(* Logix 5000 project; controller _GigaDiscovery vendor 1 type 14 code 244 rev 35.11; software revision 35.03; part 9 of 23 *)
(* tags used below, declared in another part *)
   Pylon_Sequencer : Sequencer;
   Acc_Time : REAL;   // T2 Region 2
   Auto_Cycle_Step : DINT;
   Automatic_Cycle_DB : Auto_Cycle[6];
   Cycle_Time : TIMER;
   Direction : BOOL;   // 1 = Spinta CW 0 = Spinta CCW
   Echo_HMI_Modify_Auto_Cycle_Ptr : DINT;
   Emergencies_CL1 : DINT[14];
   Gondola_Speed_Reference : DINT;
   HMI_Auto_Cycle_in_Modify : Auto_Cycle;
   HMI_Auto_Cycle_Step_Modify : DINT;
   HMI_Modify_Auto_Cycle_Ptr : DINT;
   HMI_Save_Recipe : BOOL;
   HMI_Step_in_Modify_Gondola_Speed : DINT;
   HMI_Step_in_Modify_Gondola_Time : DINT;
   HMI_Work_Auto_Cycle_Ptr : DINT;
   Jerk_Time : REAL;   // T1 Region 1
   K_Inversion : REAL;   // Fattore di Inversione
   K_Inversion_SCRV : REAL;
   LapBarsMonitor : LapBars_Monitor[41];
   LPF_WLang_Speed_to_Torq : REAL;
   ONP : DINT;   // Optional Not Present
   Oscillation_Error : REAL;
   PW_Bool : BOOL[32];
   PW_Dint : DINT[64];
   Pylon_Axe : Axe;
   Pylon_Filtered_Speed : REAL;
   RESTRAINTS_Open_Postion : BOOL[64];
   RESTRAINTS_Sector : LapBars_Sector[9];
   SCuve_K_Stop : S_Curve_Calc;
   Second_Oscillation_Done : BOOL;   // Second Oscillation End
   Start_Stop_Cycle : Sequencer;
   Stop_K_to_Zero : BOOL;
   Target_Angle : REAL;
   To_Sfty : Std_to_Sfty;
   Torque_Cmd_from_Cycle : REAL;
   TorquePos_Angle_Control : REAL;
   Work_Auto_Cycle : Auto_Cycle;
   Work_Auto_Cycle_Ptr : DINT;
(* Pylon, continued *)

ROUTINE Main   (* ladder *)
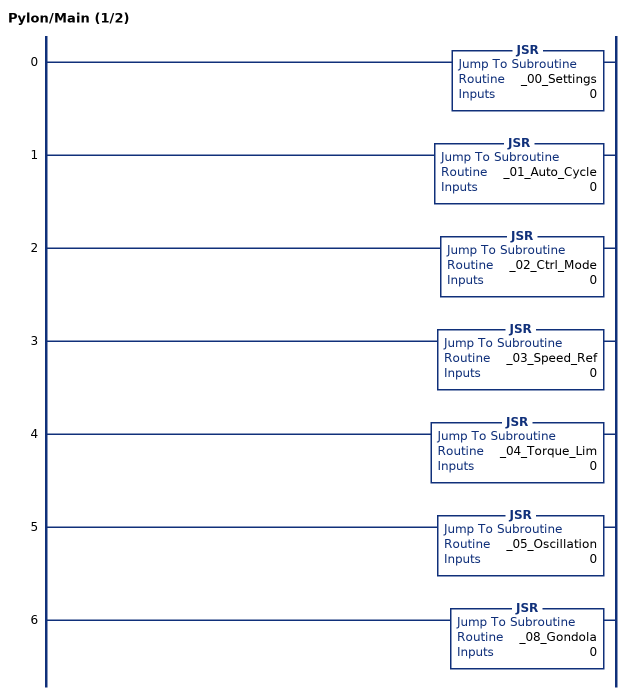
   0: JSR(_00_Settings,0);
   1: JSR(_01_Auto_Cycle,0);
   2: JSR(_02_Ctrl_Mode,0);
   3: JSR(_03_Speed_Ref,0);
   4: JSR(_04_Torque_Lim,0);
   5: JSR(_05_Oscillation,0);
   6: JSR(_08_Gondola,0);
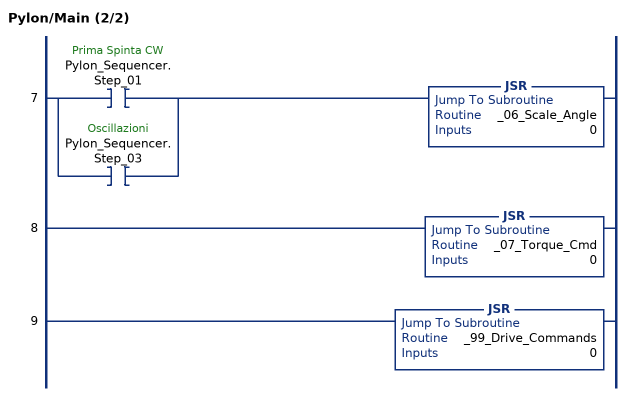
   7: [XIC(Pylon_Sequencer.Step_01) ,XIC(Pylon_Sequencer.Step_03) ]JSR(_06_Scale_Angle,0);
   8: JSR(_07_Torque_Cmd,0);
   9: JSR(_99_Drive_Commands,0);
END_ROUTINE
END_PROGRAM

PROGRAM Pylon_Oscillation   (* main routine _00_Oscillation *)
VAR
   ADD_01 : FBD_MATH := (SourceA := 0.3, SourceB := 0.5, Dest := 0.8);
   BOR_01 : FBD_BOOLEAN_OR;
   DIV_01 : FBD_MATH := (SourceA := 86.0, SourceB := 0.8, Dest := 107.5);
   DIV_02 : FBD_MATH := (SourceA := 107.5, SourceB := 0.3, Dest := 358.3333);
   GRT_01 : FBD_COMPARE;
   LES_01 : FBD_COMPARE;
   NEG_01 : FBD_MATH_ADVANCED := (Source := 77.39982, Dest := -77.39982);
   OSRI_01 : FBD_ONESHOT;
   OSRI_02 : FBD_ONESHOT;
   SCRV_01 : S_CURVE := (AccelRate := 107.5, DecelRate := 107.5, JerkRate := 358.3333, RTSTime := 1, DeltaT := 0.005);
   SCRV_02 : S_CURVE := (In := -10.0, AccelRate := 25.0, DecelRate := 25.0, JerkRate := 25.0, RTSTime := 1, Out := -10.0, DeltaT := 0.005);
   SEL_01 : SELECT := (In1 := 119.95556, In2 := 119.95556, Out := 119.95556);
   SUB_02 : FBD_MATH := (SourceA := 120.0, SourceB := 0.044444446, Dest := 119.95556);
END_VAR

ROUTINE _00_Oscillation   (* function block diagram *)
   SHEET 1
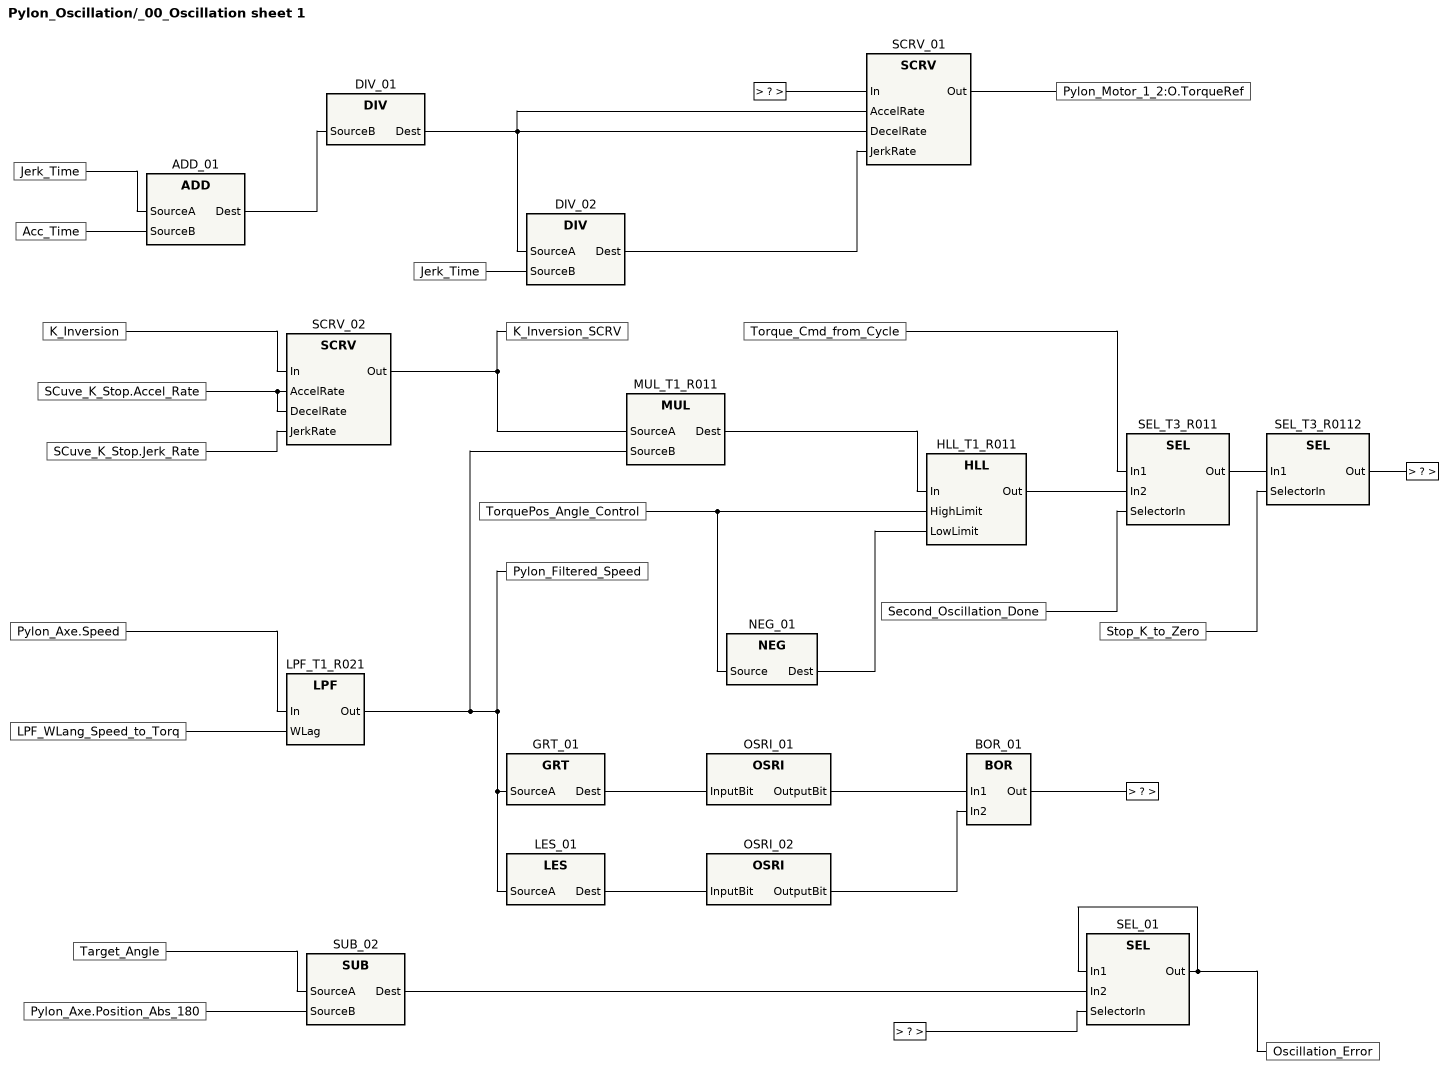
   ADD_01 : ADD(SourceA := Jerk_Time, SourceB := Acc_Time);
   SCRV_02 : SCRV(In := K_Inversion, AccelRate := SCuve_K_Stop.Accel_Rate, DecelRate := SCuve_K_Stop.Accel_Rate, JerkRate := SCuve_K_Stop.Jerk_Rate);
   LPF_T1_R021 : LPF(In := Pylon_Axe.Speed, WLag := LPF_WLang_Speed_to_Torq);
   SUB_02 : SUB(SourceA := Target_Angle, SourceB := Pylon_Axe.Position_Abs_180);
   DIV_01 : DIV(SourceB := ADD_01.Dest);
   K_Inversion_SCRV := SCRV_02.Out;
   Pylon_Filtered_Speed := LPF_T1_R021.Out;
   GRT_01 : GRT(SourceA := LPF_T1_R021.Out);
   LES_01 : LES(SourceA := LPF_T1_R021.Out);
   DIV_02 : DIV(SourceA := DIV_01.Dest, SourceB := Jerk_Time);
   MUL_T1_R011 : MUL(SourceA := SCRV_02.Out, SourceB := LPF_T1_R021.Out);
   OSRI_01 : OSRI(InputBit := GRT_01.Dest);
   OSRI_02 : OSRI(InputBit := LES_01.Dest);
   NEG_01 : NEG(Source := TorquePos_Angle_Control);
   HLL_T1_R011 : HLL(In := MUL_T1_R011.Dest, HighLimit := TorquePos_Angle_Control, LowLimit := NEG_01.Dest);
   BOR_01 : BOR(In1 := OSRI_01.OutputBit, In2 := OSRI_02.OutputBit);
   SEL_T3_R011 : SEL(In1 := Torque_Cmd_from_Cycle, In2 := HLL_T1_R011.Out, SelectorIn := Second_Oscillation_Done);
   WIRE(?) := BOR_01.Out;
   SEL_T3_R0112 : SEL(In1 := SEL_T3_R011.Out, SelectorIn := Stop_K_to_Zero);
   WIRE(?) := SEL_T3_R0112.Out;
   SCRV_01 : SCRV(In := WIRE(?), AccelRate := DIV_01.Dest, DecelRate := DIV_01.Dest, JerkRate := DIV_02.Dest);
   Pylon_Motor_1_2:O.TorqueRef := SCRV_01.Out;
   SEL_01 : SEL(In1 := SEL_01.Out, In2 := SUB_02.Dest, SelectorIn := WIRE(?));
   Oscillation_Error := SEL_01.Out;
END_ROUTINE
END_PROGRAM

PROGRAM Recipe   (* main routine Main *)
VAR
   Echo_HMI_Auto_Cycle_Step_Modify : DINT := 2;
   HMI_Cycle_Time_to_End : DINT := 145;
   Os : DINT;
   Step_Timer : TIMER := (PRE := 60000);
END_VAR

ROUTINE _01_Auto_Cycle   (* ladder *)
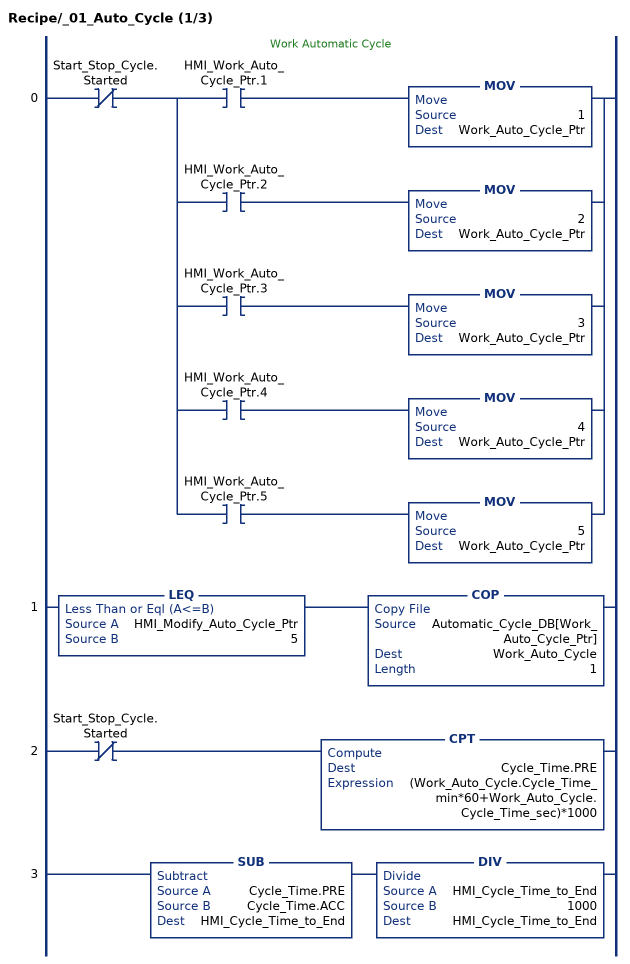
   // Work Automatic Cycle
   0: XIO(Start_Stop_Cycle.Started)[XIC(HMI_Work_Auto_Cycle_Ptr.1) MOV(1,Work_Auto_Cycle_Ptr) ,XIC(HMI_Work_Auto_Cycle_Ptr.2) MOV(2,Work_Auto_Cycle_Ptr) ,XIC(HMI_Work_Auto_Cycle_Ptr.3) MOV(3,Work_Auto_Cycle_Ptr) ,XIC(HMI_Work_Auto_Cycle_Ptr.4) MOV(4,Work_Auto_Cycle_Ptr) ,XIC(HMI_Work_Auto_Cycle_Ptr.5) MOV(5,Work_Auto_Cycle_Ptr) ];
   1: LEQ(HMI_Modify_Auto_Cycle_Ptr,5)COP(Automatic_Cycle_DB[Work_Auto_Cycle_Ptr],Work_Auto_Cycle,1);
   2: XIO(Start_Stop_Cycle.Started)CPT(Cycle_Time.PRE,(Work_Auto_Cycle.Cycle_Time_min*60+Work_Auto_Cycle.Cycle_Time_sec)*1000);
   3: SUB(Cycle_Time.PRE,Cycle_Time.ACC,HMI_Cycle_Time_to_End)DIV(HMI_Cycle_Time_to_End,1000,HMI_Cycle_Time_to_End);
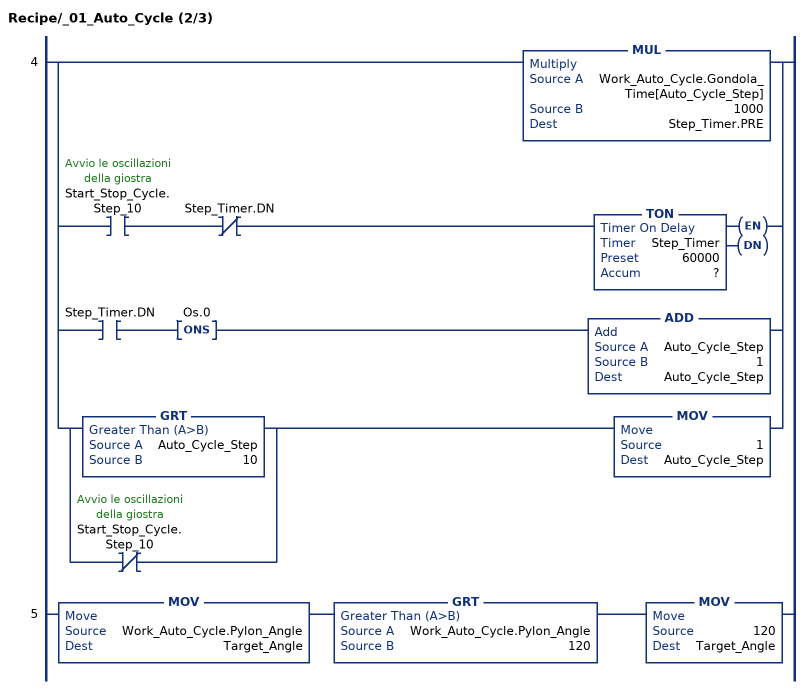
   4: [MUL(Work_Auto_Cycle.Gondola_Time[Auto_Cycle_Step],1000,Step_Timer.PRE) ,XIC(Start_Stop_Cycle.Step_10) XIO(Step_Timer.DN) TON(Step_Timer,?,?) ,XIC(Step_Timer.DN) ONS(Os.0) ADD(Auto_Cycle_Step,1,Auto_Cycle_Step) ,[GRT(Auto_Cycle_Step,10) ,XIO(Start_Stop_Cycle.Step_10) ] MOV(1,Auto_Cycle_Step) ];
   5: MOV(Work_Auto_Cycle.Pylon_Angle,Target_Angle)GRT(Work_Auto_Cycle.Pylon_Angle,120)MOV(120,Target_Angle);
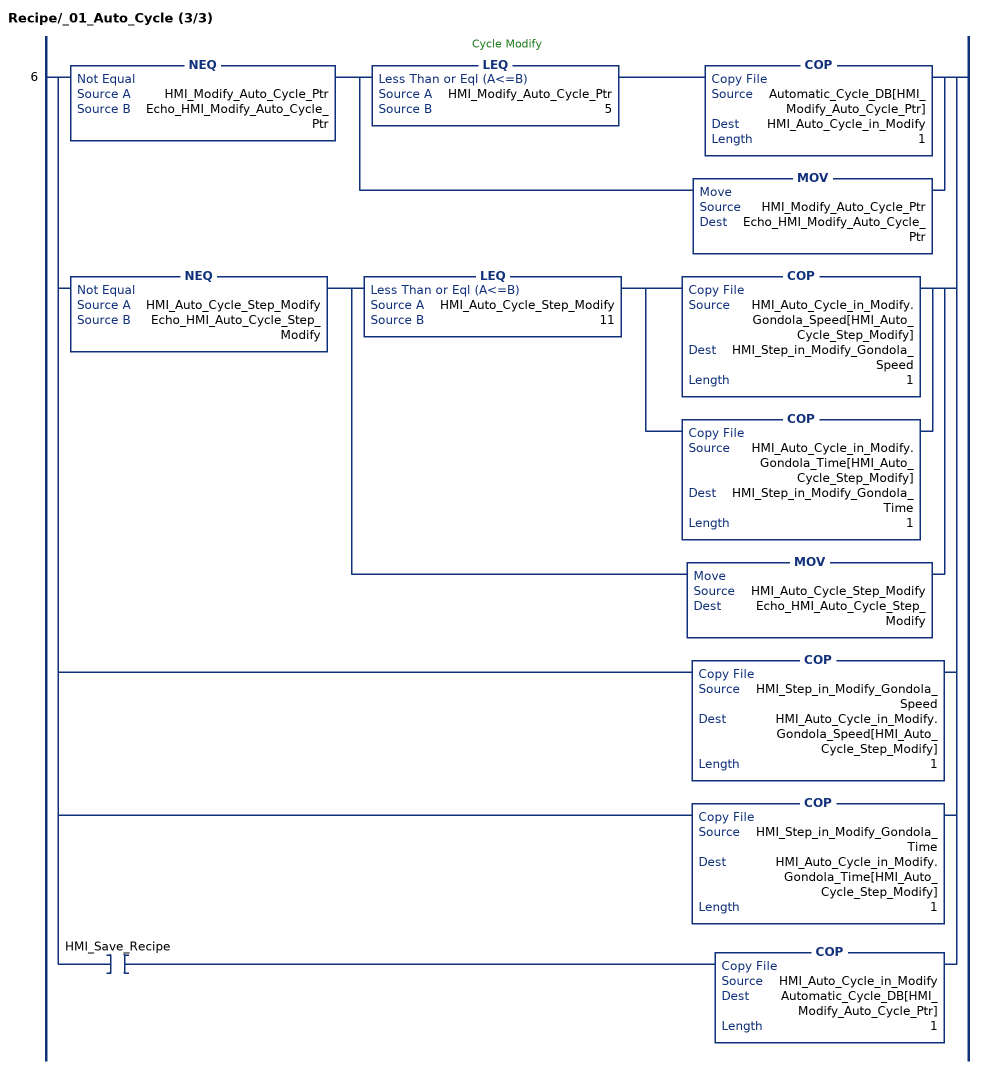
   // Cycle Modify
   6: [NEQ(HMI_Modify_Auto_Cycle_Ptr,Echo_HMI_Modify_Auto_Cycle_Ptr) [LEQ(HMI_Modify_Auto_Cycle_Ptr,5) COP(Automatic_Cycle_DB[HMI_Modify_Auto_Cycle_Ptr],HMI_Auto_Cycle_in_Modify,1) ,MOV(HMI_Modify_Auto_Cycle_Ptr,Echo_HMI_Modify_Auto_Cycle_Ptr) ] ,NEQ(HMI_Auto_Cycle_Step_Modify,Echo_HMI_Auto_Cycle_Step_Modify) [LEQ(HMI_Auto_Cycle_Step_Modify,11) [COP(HMI_Auto_Cycle_in_Modify.Gondola_Speed[HMI_Auto_Cycle_Step_Modify],HMI_Step_in_Modify_Gondola_Speed,1) ,COP(HMI_Auto_Cycle_in_Modify.Gondola_Time[HMI_Auto_Cycle_Step_Modify],HMI_Step_in_Modify_Gondola_Time,1) ] ,MOV(HMI_Auto_Cycle_Step_Modify,Echo_HMI_Auto_Cycle_Step_Modify) ] ,[COP(HMI_Step_in_Modify_Gondola_Speed,HMI_Auto_Cycle_in_Modify.Gondola_Speed[HMI_Auto_Cycle_Step_Modify],1) ,COP(HMI_Step_in_Modify_Gondola_Time,HMI_Auto_Cycle_in_Modify.Gondola_Time[HMI_Auto_Cycle_Step_Modify],1) ] ,XIC(HMI_Save_Recipe) COP(HMI_Auto_Cycle_in_Modify,Automatic_Cycle_DB[HMI_Modify_Auto_Cycle_Ptr],1) ];
END_ROUTINE

ROUTINE _02_Maintenance   (* ladder *)
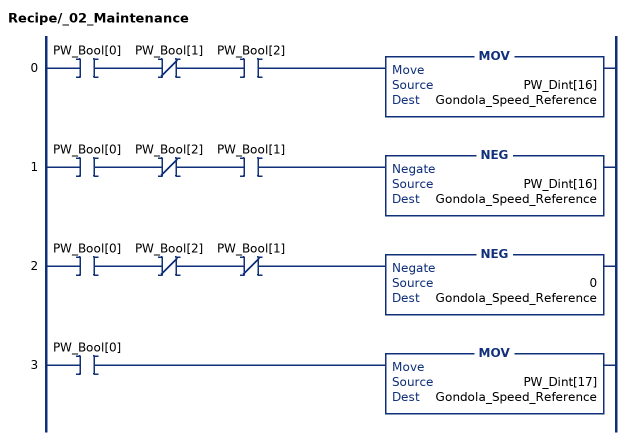
   0: XIC(PW_Bool[0])XIO(PW_Bool[1])XIC(PW_Bool[2])MOV(PW_Dint[16],Gondola_Speed_Reference);
   1: XIC(PW_Bool[0])XIO(PW_Bool[2])XIC(PW_Bool[1])NEG(PW_Dint[16],Gondola_Speed_Reference);
   2: XIC(PW_Bool[0])XIO(PW_Bool[2])XIO(PW_Bool[1])NEG(0,Gondola_Speed_Reference);
   3: XIC(PW_Bool[0])MOV(PW_Dint[17],Gondola_Speed_Reference);
END_ROUTINE

ROUTINE Main   (* ladder *)
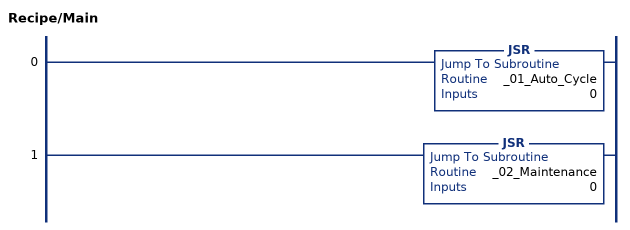
   0: JSR(_01_Auto_Cycle,0);
   1: JSR(_02_Maintenance,0);
END_ROUTINE
END_PROGRAM

PROGRAM Restraints   (* main routine Main *)
VAR
   ADD_02 : FBD_MATH := (SourceA := -11.0, SourceB := 11.0);
   DIV_01 : FBD_MATH := (SourceB := 100.0);
   In_FGEN_01 : FUNCTION_GENERATOR := (XY1Size := 2, Out := 0.0061035156);
   In_FGEN_02 : FUNCTION_GENERATOR := (XY1Size := 2);
   In_FGEN_03 : FUNCTION_GENERATOR := (In := -2.125, XY1Size := 2, Out := -0.025939941);
   In_FGEN_04 : FUNCTION_GENERATOR := (XY1Size := 2);
   In_FGEN_05 : FUNCTION_GENERATOR := (In := -2.0625, XY1Size := 2, Out := -0.025177002);
   In_FGEN_06 : FUNCTION_GENERATOR := (XY1Size := 2);
   In_FGEN_07 : FUNCTION_GENERATOR := (In := -2.25, XY1Size := 2, Out := -0.02746582);
   In_FGEN_08 : FUNCTION_GENERATOR := (XY1Size := 2);
   LapBarsGeneral_Monitor : BOOL := 1; {access Read Only}
   LPF_01 : FILTER_LOW_PASS := (WLag := 1.7453293, Order := 1, RTSTime := 1, DeltaT := 0.001);
   LPF_02 : FILTER_LOW_PASS := (WLag := 0.34906584, Order := 1, RTSTime := 1, DeltaT := 0.001);
   LPF_04 : FILTER_LOW_PASS := (In := -0.025939941, Order := 1, RTSTime := 1, Out := -0.02593994, DeltaT := 0.001, Status := 16#0000_0003, InstructFault := 1, WLagInv := 1);
   LPF_05 : FILTER_LOW_PASS := (WLag := 2.0, Order := 2, RTSTime := 1, DeltaT := 0.001);
   Ptr_LapBars : DINT := 33; {access Read Only}
   RAD_01 : FBD_MATH_ADVANCED := (Source := 100.0, Dest := 1.7453293);
   RAD_02 : FBD_MATH_ADVANCED := (Source := 20.0, Dest := 0.34906584);
   Seat_Auxiliary_Ch_Memory : INT := -1;
END_VAR

ROUTINE _01_Memory   (* structured text *)
   if Start_Stop_Cycle.Step_00 then
   	for Ptr_LapBars :=1 to 40 do
   		if RESTRAINTS_Open_Postion[Ptr_LapBars] then
   			LapBarsMonitor[Ptr_LapBars].Sensor_Open_Memory := 1;
   		end_if;
   	end_for;
   end_if;
   
   if Start_Stop_Cycle.Step_01 then
   	for Ptr_LapBars :=1 to 40 do
   		LapBarsMonitor[Ptr_LapBars].Sensor_Open_Memory := 0;
   	end_for;
   end_if;
   
   LapBarsGeneral_Monitor := 0;
   for Ptr_LapBars :=1 to 40 do
   	LapBarsMonitor[Ptr_LapBars].Status := 0;
   	if 	LapBarsMonitor[Ptr_LapBars].Sensor_Open_Memory then
   		LapBarsMonitor[Ptr_LapBars].Status := 1;
   		LapBarsGeneral_Monitor := 1;
   	end_if;
   end_for;
   for Ptr_LapBars :=1 to 8 do
   	if RESTRAINTS_Sector[Ptr_LapBars].I_Close_Position.O1 then
   	else
   		LapBarsMonitor[Ptr_LapBars].Status := 1;
   		LapBarsGeneral_Monitor := 1;
   	end_if;
   end_for;
   
END_ROUTINE

ROUTINE _02_Seats_Memory   (* ladder *)
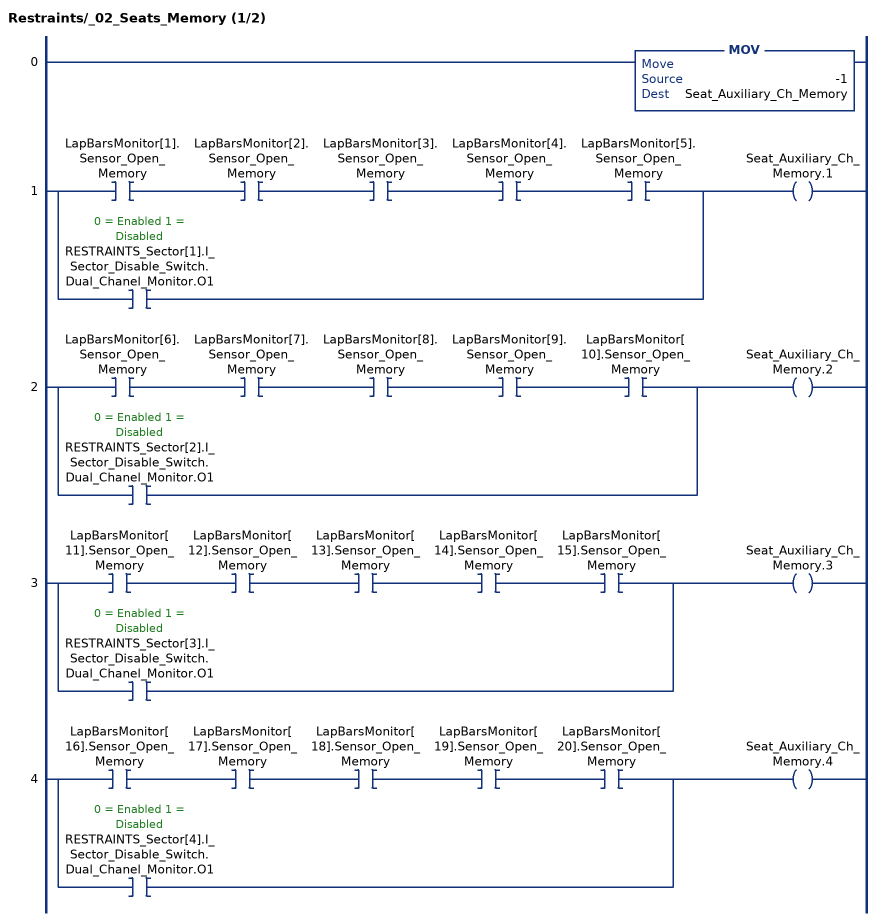
   0: MOV(-1,Seat_Auxiliary_Ch_Memory);
   1: [XIC(LapBarsMonitor[1].Sensor_Open_Memory) XIC(LapBarsMonitor[2].Sensor_Open_Memory) XIC(LapBarsMonitor[3].Sensor_Open_Memory) XIC(LapBarsMonitor[4].Sensor_Open_Memory) XIC(LapBarsMonitor[5].Sensor_Open_Memory) ,XIC(RESTRAINTS_Sector[1].I_Sector_Disable_Switch.Dual_Chanel_Monitor.O1) ]OTE(Seat_Auxiliary_Ch_Memory.1);
   2: [XIC(LapBarsMonitor[6].Sensor_Open_Memory) XIC(LapBarsMonitor[7].Sensor_Open_Memory) XIC(LapBarsMonitor[8].Sensor_Open_Memory) XIC(LapBarsMonitor[9].Sensor_Open_Memory) XIC(LapBarsMonitor[10].Sensor_Open_Memory) ,XIC(RESTRAINTS_Sector[2].I_Sector_Disable_Switch.Dual_Chanel_Monitor.O1) ]OTE(Seat_Auxiliary_Ch_Memory.2);
   3: [XIC(LapBarsMonitor[11].Sensor_Open_Memory) XIC(LapBarsMonitor[12].Sensor_Open_Memory) XIC(LapBarsMonitor[13].Sensor_Open_Memory) XIC(LapBarsMonitor[14].Sensor_Open_Memory) XIC(LapBarsMonitor[15].Sensor_Open_Memory) ,XIC(RESTRAINTS_Sector[3].I_Sector_Disable_Switch.Dual_Chanel_Monitor.O1) ]OTE(Seat_Auxiliary_Ch_Memory.3);
   4: [XIC(LapBarsMonitor[16].Sensor_Open_Memory) XIC(LapBarsMonitor[17].Sensor_Open_Memory) XIC(LapBarsMonitor[18].Sensor_Open_Memory) XIC(LapBarsMonitor[19].Sensor_Open_Memory) XIC(LapBarsMonitor[20].Sensor_Open_Memory) ,XIC(RESTRAINTS_Sector[4].I_Sector_Disable_Switch.Dual_Chanel_Monitor.O1) ]OTE(Seat_Auxiliary_Ch_Memory.4);
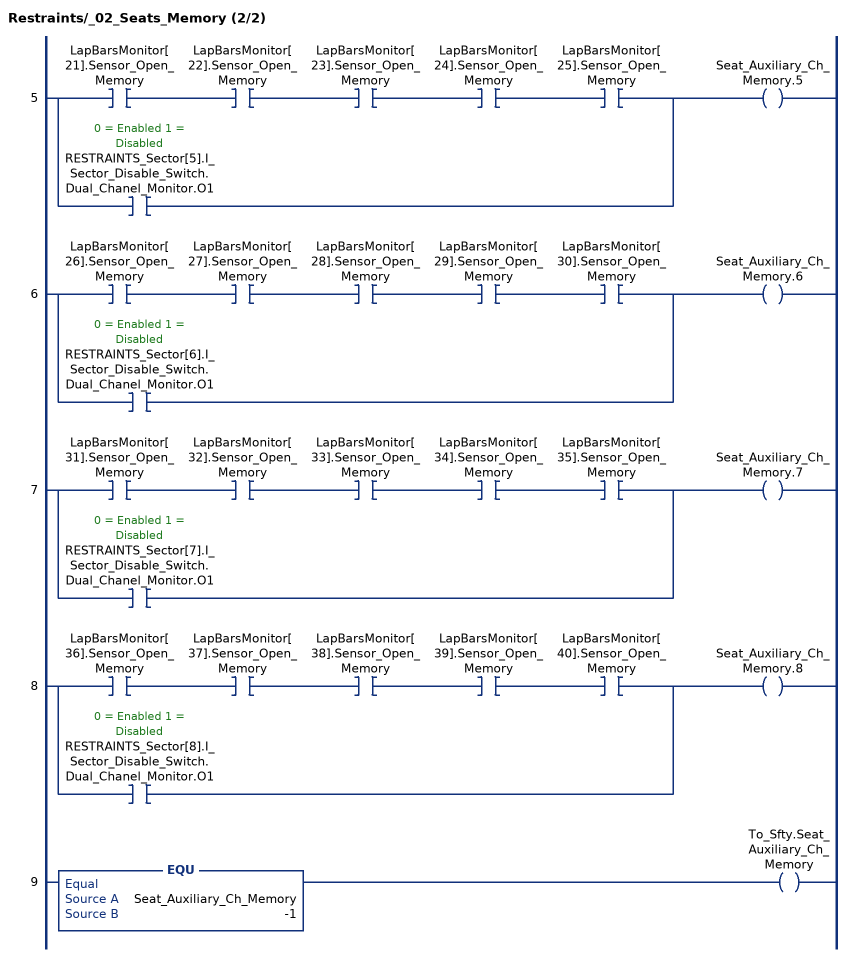
   5: [XIC(LapBarsMonitor[21].Sensor_Open_Memory) XIC(LapBarsMonitor[22].Sensor_Open_Memory) XIC(LapBarsMonitor[23].Sensor_Open_Memory) XIC(LapBarsMonitor[24].Sensor_Open_Memory) XIC(LapBarsMonitor[25].Sensor_Open_Memory) ,XIC(RESTRAINTS_Sector[5].I_Sector_Disable_Switch.Dual_Chanel_Monitor.O1) ]OTE(Seat_Auxiliary_Ch_Memory.5);
   6: [XIC(LapBarsMonitor[26].Sensor_Open_Memory) XIC(LapBarsMonitor[27].Sensor_Open_Memory) XIC(LapBarsMonitor[28].Sensor_Open_Memory) XIC(LapBarsMonitor[29].Sensor_Open_Memory) XIC(LapBarsMonitor[30].Sensor_Open_Memory) ,XIC(RESTRAINTS_Sector[6].I_Sector_Disable_Switch.Dual_Chanel_Monitor.O1) ]OTE(Seat_Auxiliary_Ch_Memory.6);
   7: [XIC(LapBarsMonitor[31].Sensor_Open_Memory) XIC(LapBarsMonitor[32].Sensor_Open_Memory) XIC(LapBarsMonitor[33].Sensor_Open_Memory) XIC(LapBarsMonitor[34].Sensor_Open_Memory) XIC(LapBarsMonitor[35].Sensor_Open_Memory) ,XIC(RESTRAINTS_Sector[7].I_Sector_Disable_Switch.Dual_Chanel_Monitor.O1) ]OTE(Seat_Auxiliary_Ch_Memory.7);
   8: [XIC(LapBarsMonitor[36].Sensor_Open_Memory) XIC(LapBarsMonitor[37].Sensor_Open_Memory) XIC(LapBarsMonitor[38].Sensor_Open_Memory) XIC(LapBarsMonitor[39].Sensor_Open_Memory) XIC(LapBarsMonitor[40].Sensor_Open_Memory) ,XIC(RESTRAINTS_Sector[8].I_Sector_Disable_Switch.Dual_Chanel_Monitor.O1) ]OTE(Seat_Auxiliary_Ch_Memory.8);